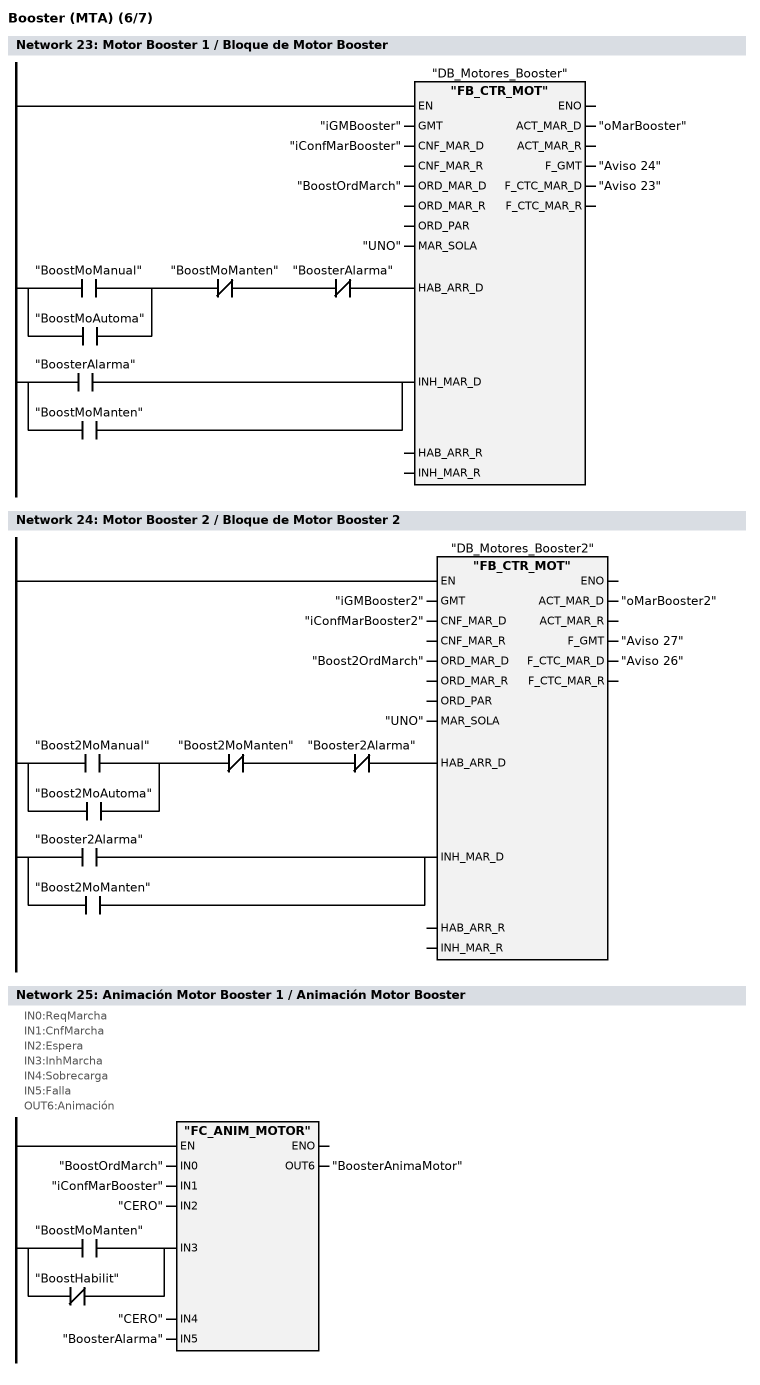
   RUNG wire#powerrail
      "DB_Motores_Booster"(HAB_ARR_D := wire#w2, INH_MAR_D := wire#w3, GMT := "iGMBooster", CNF_MAR_D := "iConfMarBooster", CNF_MAR_R :=, ORD_MAR_D := "BoostOrdMarch", ORD_MAR_R :=, ORD_PAR :=, MAR_SOLA := "UNO", HAB_ARR_R :=, INH_MAR_R :=, ACT_MAR_D => "oMarBooster", ACT_MAR_R =>, F_GMT => "Aviso 24", F_CTC_MAR_D => "Aviso 23", F_CTC_MAR_R =>)
   END_RUNG
   RUNG wire#powerrail
      Contact( "BoostMoManual" )
      wire#w1
      I_Contact( "BoostMoManten" )
      I_Contact( "BoosterAlarma" )
   END_RUNG wire#w2
   RUNG wire#powerrail
      Contact( "BoostMoAutoma" )
   END_RUNG wire#w1
   RUNG wire#powerrail
      Contact( "BoosterAlarma" )
   END_RUNG wire#w3
   RUNG wire#powerrail
      Contact( "BoostMoManten" )
   END_RUNG wire#w3
   // the same network as SCL:
   "DB_Motores_Booster"(GMT := "iGMBooster",   // "FB_CTR_MOT"
                        CNF_MAR_D := "iConfMarBooster",
                        ORD_MAR_D := "BoostOrdMarch",
                        MAR_SOLA := "UNO",
                        HAB_ARR_D := ("BoostMoManual" OR "BoostMoAutoma") AND NOT "BoostMoManten" AND NOT "BoosterAlarma",
                        INH_MAR_D := "BoosterAlarma" OR "BoostMoManten",
                        ACT_MAR_D => "oMarBooster",
                        F_GMT => "Aviso 24",
                        F_CTC_MAR_D => "Aviso 23");
END_REGION

REGION Network 24: Motor Booster 2 / Bloque de Motor Booster 2
   RUNG wire#powerrail
      "DB_Motores_Booster2"(HAB_ARR_D := wire#w2, INH_MAR_D := wire#w3, GMT := "iGMBooster2", CNF_MAR_D := "iConfMarBooster2", CNF_MAR_R :=, ORD_MAR_D := "Boost2OrdMarch", ORD_MAR_R :=, ORD_PAR :=, MAR_SOLA := "UNO", HAB_ARR_R :=, INH_MAR_R :=, ACT_MAR_D => "oMarBooster2", ACT_MAR_R =>, F_GMT => "Aviso 27", F_CTC_MAR_D => "Aviso 26", F_CTC_MAR_R =>)
   END_RUNG
   RUNG wire#powerrail
      Contact( "Boost2MoManual" )
      wire#w1
      I_Contact( "Boost2MoManten" )
      I_Contact( "Booster2Alarma" )
   END_RUNG wire#w2
   RUNG wire#powerrail
      Contact( "Boost2MoAutoma" )
   END_RUNG wire#w1
   RUNG wire#powerrail
      Contact( "Booster2Alarma" )
   END_RUNG wire#w3
   RUNG wire#powerrail
      Contact( "Boost2MoManten" )
   END_RUNG wire#w3
   // the same network as SCL:
   "DB_Motores_Booster2"(GMT := "iGMBooster2",   // "FB_CTR_MOT"
                         CNF_MAR_D := "iConfMarBooster2",
                         ORD_MAR_D := "Boost2OrdMarch",
                         MAR_SOLA := "UNO",
                         HAB_ARR_D := ("Boost2MoManual" OR "Boost2MoAutoma") AND NOT "Boost2MoManten" AND NOT "Booster2Alarma",
                         INH_MAR_D := "Booster2Alarma" OR "Boost2MoManten",
                         ACT_MAR_D => "oMarBooster2",
                         F_GMT => "Aviso 27",
                         F_CTC_MAR_D => "Aviso 26");
END_REGION

REGION Network 25: Animación Motor Booster 1 / Animación Motor Booster
   // IN0:ReqMarcha
   // IN1:CnfMarcha
   // IN2:Espera
   // IN3:InhMarcha
   // IN4:Sobrecarga
   // IN5:Falla
   // OUT6:Animación
   RUNG wire#powerrail
      "FC_ANIM_MOTOR"(IN0 := "BoostOrdMarch", IN1 := "iConfMarBooster", IN2 := "CERO", IN3 := wire#w1, IN4 := "CERO", IN5 := "BoosterAlarma", OUT6 => "BoosterAnimaMotor")
   END_RUNG
   RUNG wire#powerrail
      Contact( "BoostMoManten" )
   END_RUNG wire#w1
   RUNG wire#powerrail
      I_Contact( "BoostHabilit" )
   END_RUNG wire#w1
   // the same network as SCL:
   "FC_ANIM_MOTOR"(IN0 := "BoostOrdMarch",
                   IN1 := "iConfMarBooster",
                   IN2 := "CERO",
                   IN3 := "BoostMoManten" OR NOT "BoostHabilit",
                   IN4 := "CERO",
                   IN5 := "BoosterAlarma",
                   OUT6 => "BoosterAnimaMotor");
END_REGION

REGION Network 26: Animación Motor Booster 2
   // IN0:ReqMarcha
   // IN1:CnfMarcha
   // IN2:Espera
   // IN3:InhMarcha
   // IN4:Sobrecarga
   // IN5:Falla
   // OUT6:Animación
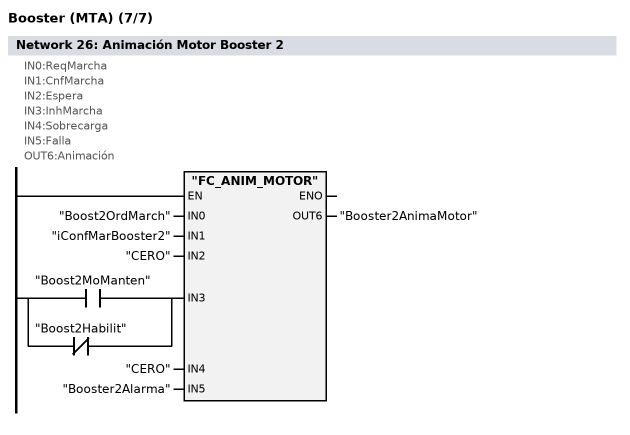
   RUNG wire#powerrail
      "FC_ANIM_MOTOR"(IN0 := "Boost2OrdMarch", IN1 := "iConfMarBooster2", IN2 := "CERO", IN3 := wire#w1, IN4 := "CERO", IN5 := "Booster2Alarma", OUT6 => "Booster2AnimaMotor")
   END_RUNG
   RUNG wire#powerrail
      Contact( "Boost2MoManten" )
   END_RUNG wire#w1
   RUNG wire#powerrail
      I_Contact( "Boost2Habilit" )
   END_RUNG wire#w1
   // the same network as SCL:
   "FC_ANIM_MOTOR"(IN0 := "Boost2OrdMarch",
                   IN1 := "iConfMarBooster2",
                   IN2 := "CERO",
                   IN3 := "Boost2MoManten" OR NOT "Boost2Habilit",
                   IN4 := "CERO",
                   IN5 := "Booster2Alarma",
                   OUT6 => "Booster2AnimaMotor");
END_REGION
END_FUNCTION

// folder: Compresores/Alta

FUNCTION "CompresoresAltaMTA" : Void   // FC13, LAD
{ S7_Optimized_Access := 'FALSE' }
VERSION : 0.1
BEGIN

REGION Network 1
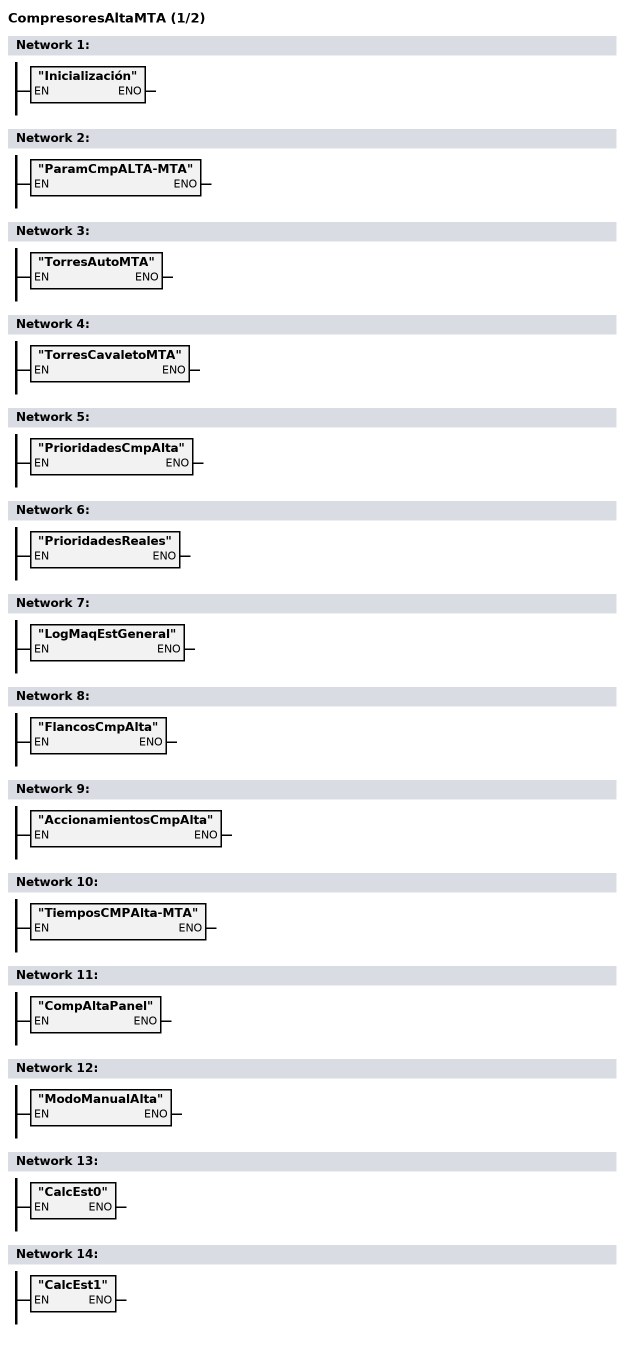
   RUNG wire#powerrail
      "Inicialización"()
   END_RUNG
   // the same network as SCL:
   "Inicialización"();
END_REGION

REGION Network 2
   RUNG wire#powerrail
      "ParamCmpALTA-MTA"()
   END_RUNG
   // the same network as SCL:
   "ParamCmpALTA-MTA"();
END_REGION

REGION Network 3
   RUNG wire#powerrail
      "TorresAutoMTA"()
   END_RUNG
   // the same network as SCL:
   "TorresAutoMTA"();
END_REGION

REGION Network 4
   RUNG wire#powerrail
      "TorresCavaletoMTA"()
   END_RUNG
   // the same network as SCL:
   "TorresCavaletoMTA"();
END_REGION

REGION Network 5
   RUNG wire#powerrail
      "PrioridadesCmpAlta"()
   END_RUNG
   // the same network as SCL:
   "PrioridadesCmpAlta"();
END_REGION

REGION Network 6
   RUNG wire#powerrail
      "PrioridadesReales"()
   END_RUNG
   // the same network as SCL:
   "PrioridadesReales"();
END_REGION

REGION Network 7
   RUNG wire#powerrail
      "LogMaqEstGeneral"()
   END_RUNG
   // the same network as SCL:
   "LogMaqEstGeneral"();
END_REGION

REGION Network 8
   RUNG wire#powerrail
      "FlancosCmpAlta"()
   END_RUNG
   // the same network as SCL:
   "FlancosCmpAlta"();
END_REGION

REGION Network 9
   RUNG wire#powerrail
      "AccionamientosCmpAlta"()
   END_RUNG
   // the same network as SCL:
   "AccionamientosCmpAlta"();
END_REGION

REGION Network 10
   RUNG wire#powerrail
      "TiemposCMPAlta-MTA"()
   END_RUNG
   // the same network as SCL:
   "TiemposCMPAlta-MTA"();
END_REGION

REGION Network 11
   RUNG wire#powerrail
      "CompAltaPanel"()
   END_RUNG
   // the same network as SCL:
   "CompAltaPanel"();
END_REGION

REGION Network 12
   RUNG wire#powerrail
      "ModoManualAlta"()
   END_RUNG
   // the same network as SCL:
   "ModoManualAlta"();
END_REGION

REGION Network 13
   RUNG wire#powerrail
      "CalcEst0"()
   END_RUNG
   // the same network as SCL:
   "CalcEst0"();
END_REGION

REGION Network 14
   RUNG wire#powerrail
      "CalcEst1"()
   END_RUNG
   // the same network as SCL:
   "CalcEst1"();
END_REGION

REGION Network 15
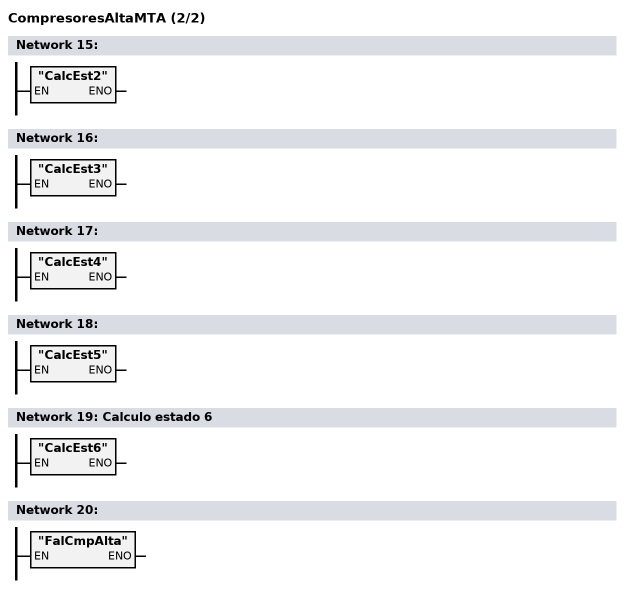
   RUNG wire#powerrail
      "CalcEst2"()
   END_RUNG
   // the same network as SCL:
   "CalcEst2"();
END_REGION

REGION Network 16
   RUNG wire#powerrail
      "CalcEst3"()
   END_RUNG
   // the same network as SCL:
   "CalcEst3"();
END_REGION

REGION Network 17
   RUNG wire#powerrail
      "CalcEst4"()
   END_RUNG
   // the same network as SCL:
   "CalcEst4"();
END_REGION

REGION Network 18
   RUNG wire#powerrail
      "CalcEst5"()
   END_RUNG
   // the same network as SCL:
   "CalcEst5"();
END_REGION

REGION Network 19: Calculo estado 6
   RUNG wire#powerrail
      "CalcEst6"()
   END_RUNG
   // the same network as SCL:
   "CalcEst6"();
END_REGION

REGION Network 20
   RUNG wire#powerrail
      "FalCmpAlta"()
   END_RUNG
   // the same network as SCL:
   "FalCmpAlta"();
END_REGION
END_FUNCTION

FUNCTION "ParamCmpALTA-MTA" : Void   // FC30, LAD
{ S7_Optimized_Access := 'FALSE' }
VERSION : 0.1
BEGIN

REGION Network 1
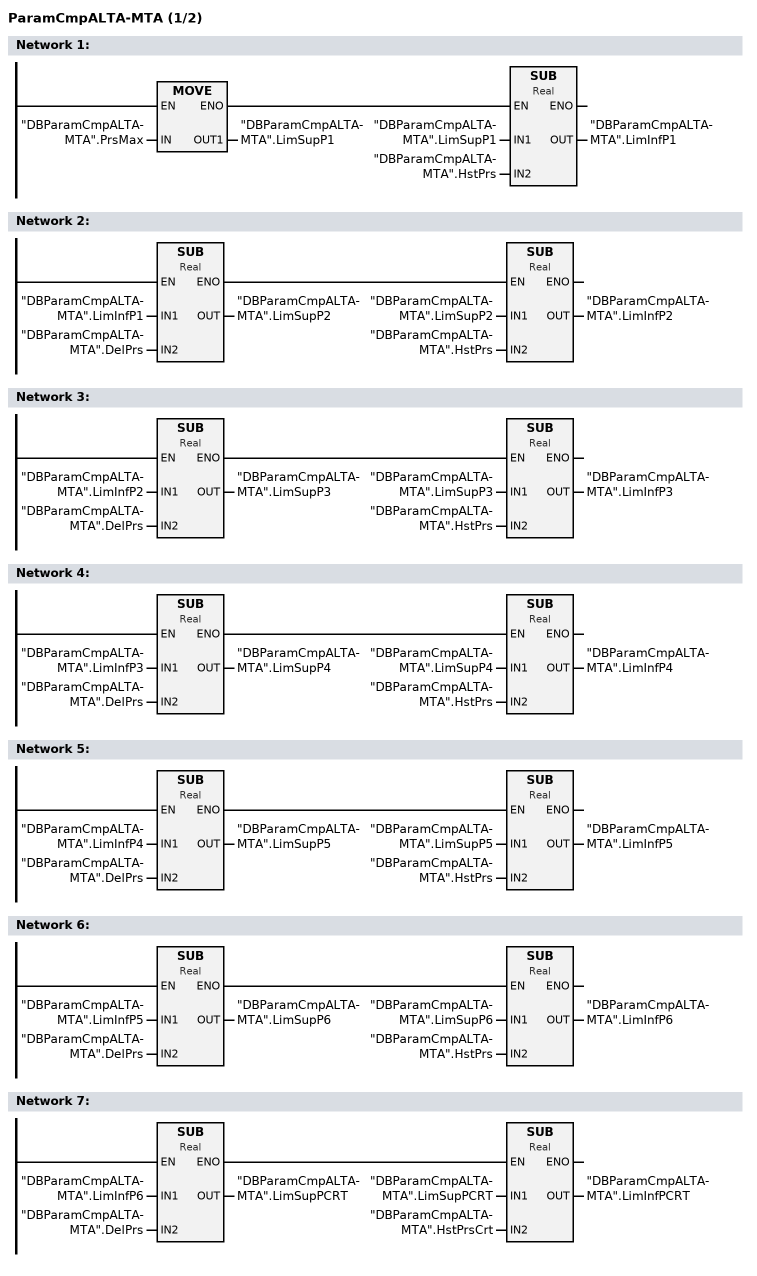
   RUNG wire#powerrail
      { S7_GenerateENO := "TRUE" } Move(in := "DBParamCmpALTA-MTA".PrsMax, out1 => "DBParamCmpALTA-MTA".LimSupP1)
      { S7_Templates := "SrcType := Real"; S7_GenerateENO := "TRUE" } Sub(in1 := "DBParamCmpALTA-MTA".LimSupP1, in2 := "DBParamCmpALTA-MTA".HstPrs, out => "DBParamCmpALTA-MTA".LimInfP1)
   END_RUNG
   // the same network as SCL:
   // ENO of a box is taken as its EN; it also drops when the box reports an error
   "DBParamCmpALTA-MTA".LimSupP1 := "DBParamCmpALTA-MTA".PrsMax;
   "DBParamCmpALTA-MTA".LimInfP1 := "DBParamCmpALTA-MTA".LimSupP1 - "DBParamCmpALTA-MTA".HstPrs;
END_REGION

REGION Network 2
   RUNG wire#powerrail
      { S7_Templates := "SrcType := Real"; S7_GenerateENO := "TRUE" } Sub(in1 := "DBParamCmpALTA-MTA".LimInfP1, in2 := "DBParamCmpALTA-MTA".DelPrs, out => "DBParamCmpALTA-MTA".LimSupP2)
      { S7_Templates := "SrcType := Real"; S7_GenerateENO := "TRUE" } Sub(in1 := "DBParamCmpALTA-MTA".LimSupP2, in2 := "DBParamCmpALTA-MTA".HstPrs, out => "DBParamCmpALTA-MTA".LimInfP2)
   END_RUNG
   // the same network as SCL:
   // ENO of a box is taken as its EN; it also drops when the box reports an error
   "DBParamCmpALTA-MTA".LimSupP2 := "DBParamCmpALTA-MTA".LimInfP1 - "DBParamCmpALTA-MTA".DelPrs;
   "DBParamCmpALTA-MTA".LimInfP2 := "DBParamCmpALTA-MTA".LimSupP2 - "DBParamCmpALTA-MTA".HstPrs;
END_REGION

REGION Network 3
   RUNG wire#powerrail
      { S7_Templates := "SrcType := Real"; S7_GenerateENO := "TRUE" } Sub(in1 := "DBParamCmpALTA-MTA".LimInfP2, in2 := "DBParamCmpALTA-MTA".DelPrs, out => "DBParamCmpALTA-MTA".LimSupP3)
      { S7_Templates := "SrcType := Real"; S7_GenerateENO := "TRUE" } Sub(in1 := "DBParamCmpALTA-MTA".LimSupP3, in2 := "DBParamCmpALTA-MTA".HstPrs, out => "DBParamCmpALTA-MTA".LimInfP3)
   END_RUNG
   // the same network as SCL:
   // ENO of a box is taken as its EN; it also drops when the box reports an error
   "DBParamCmpALTA-MTA".LimSupP3 := "DBParamCmpALTA-MTA".LimInfP2 - "DBParamCmpALTA-MTA".DelPrs;
   "DBParamCmpALTA-MTA".LimInfP3 := "DBParamCmpALTA-MTA".LimSupP3 - "DBParamCmpALTA-MTA".HstPrs;
END_REGION

REGION Network 4
   RUNG wire#powerrail
      { S7_Templates := "SrcType := Real"; S7_GenerateENO := "TRUE" } Sub(in1 := "DBParamCmpALTA-MTA".LimInfP3, in2 := "DBParamCmpALTA-MTA".DelPrs, out => "DBParamCmpALTA-MTA".LimSupP4)
      { S7_Templates := "SrcType := Real"; S7_GenerateENO := "TRUE" } Sub(in1 := "DBParamCmpALTA-MTA".LimSupP4, in2 := "DBParamCmpALTA-MTA".HstPrs, out => "DBParamCmpALTA-MTA".LimInfP4)
   END_RUNG
   // the same network as SCL:
   // ENO of a box is taken as its EN; it also drops when the box reports an error
   "DBParamCmpALTA-MTA".LimSupP4 := "DBParamCmpALTA-MTA".LimInfP3 - "DBParamCmpALTA-MTA".DelPrs;
   "DBParamCmpALTA-MTA".LimInfP4 := "DBParamCmpALTA-MTA".LimSupP4 - "DBParamCmpALTA-MTA".HstPrs;
END_REGION

REGION Network 5
   RUNG wire#powerrail
      { S7_Templates := "SrcType := Real"; S7_GenerateENO := "TRUE" } Sub(in1 := "DBParamCmpALTA-MTA".LimInfP4, in2 := "DBParamCmpALTA-MTA".DelPrs, out => "DBParamCmpALTA-MTA".LimSupP5)
      { S7_Templates := "SrcType := Real"; S7_GenerateENO := "TRUE" } Sub(in1 := "DBParamCmpALTA-MTA".LimSupP5, in2 := "DBParamCmpALTA-MTA".HstPrs, out => "DBParamCmpALTA-MTA".LimInfP5)
   END_RUNG
   // the same network as SCL:
   // ENO of a box is taken as its EN; it also drops when the box reports an error
   "DBParamCmpALTA-MTA".LimSupP5 := "DBParamCmpALTA-MTA".LimInfP4 - "DBParamCmpALTA-MTA".DelPrs;
   "DBParamCmpALTA-MTA".LimInfP5 := "DBParamCmpALTA-MTA".LimSupP5 - "DBParamCmpALTA-MTA".HstPrs;
END_REGION

REGION Network 6
   RUNG wire#powerrail
      { S7_Templates := "SrcType := Real"; S7_GenerateENO := "TRUE" } Sub(in1 := "DBParamCmpALTA-MTA".LimInfP5, in2 := "DBParamCmpALTA-MTA".DelPrs, out => "DBParamCmpALTA-MTA".LimSupP6)
      { S7_Templates := "SrcType := Real"; S7_GenerateENO := "TRUE" } Sub(in1 := "DBParamCmpALTA-MTA".LimSupP6, in2 := "DBParamCmpALTA-MTA".HstPrs, out => "DBParamCmpALTA-MTA".LimInfP6)
   END_RUNG
   // the same network as SCL:
   // ENO of a box is taken as its EN; it also drops when the box reports an error
   "DBParamCmpALTA-MTA".LimSupP6 := "DBParamCmpALTA-MTA".LimInfP5 - "DBParamCmpALTA-MTA".DelPrs;
   "DBParamCmpALTA-MTA".LimInfP6 := "DBParamCmpALTA-MTA".LimSupP6 - "DBParamCmpALTA-MTA".HstPrs;
END_REGION

REGION Network 7
   RUNG wire#powerrail
      { S7_Templates := "SrcType := Real"; S7_GenerateENO := "TRUE" } Sub(in1 := "DBParamCmpALTA-MTA".LimInfP6, in2 := "DBParamCmpALTA-MTA".DelPrs, out => "DBParamCmpALTA-MTA".LimSupPCRT)
      { S7_Templates := "SrcType := Real"; S7_GenerateENO := "TRUE" } Sub(in1 := "DBParamCmpALTA-MTA".LimSupPCRT, in2 := "DBParamCmpALTA-MTA".HstPrsCrt, out => "DBParamCmpALTA-MTA".LimInfPCRT)
   END_RUNG
   // the same network as SCL:
   // ENO of a box is taken as its EN; it also drops when the box reports an error
   "DBParamCmpALTA-MTA".LimSupPCRT := "DBParamCmpALTA-MTA".LimInfP6 - "DBParamCmpALTA-MTA".DelPrs;
   "DBParamCmpALTA-MTA".LimInfPCRT := "DBParamCmpALTA-MTA".LimSupPCRT - "DBParamCmpALTA-MTA".HstPrsCrt;
END_REGION

REGION Network 8: Falla General Flujostato Cavaleto
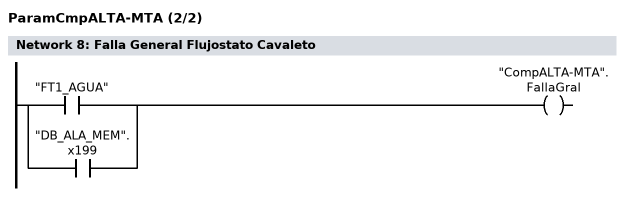
   RUNG wire#powerrail
      Contact( "FT1_AGUA" )
      wire#w1
      Coil( "CompALTA-MTA".FallaGral )
   END_RUNG
   RUNG wire#powerrail
      Contact( "DB_ALA_MEM".x199 )
   END_RUNG wire#w1
   // the same network as SCL:
   "CompALTA-MTA".FallaGral := "FT1_AGUA" OR "DB_ALA_MEM".x199;
END_REGION
END_FUNCTION

FUNCTION "TiemposCMPAlta-MTA" : Void   // FC31, LAD
{ S7_Optimized_Access := 'FALSE' }
VERSION : 0.1
   VAR_TEMP   // added for the SCL form of the ladder/FBD networks
      _s5time1 : S5Time;
   END_VAR
BEGIN

REGION Network 1
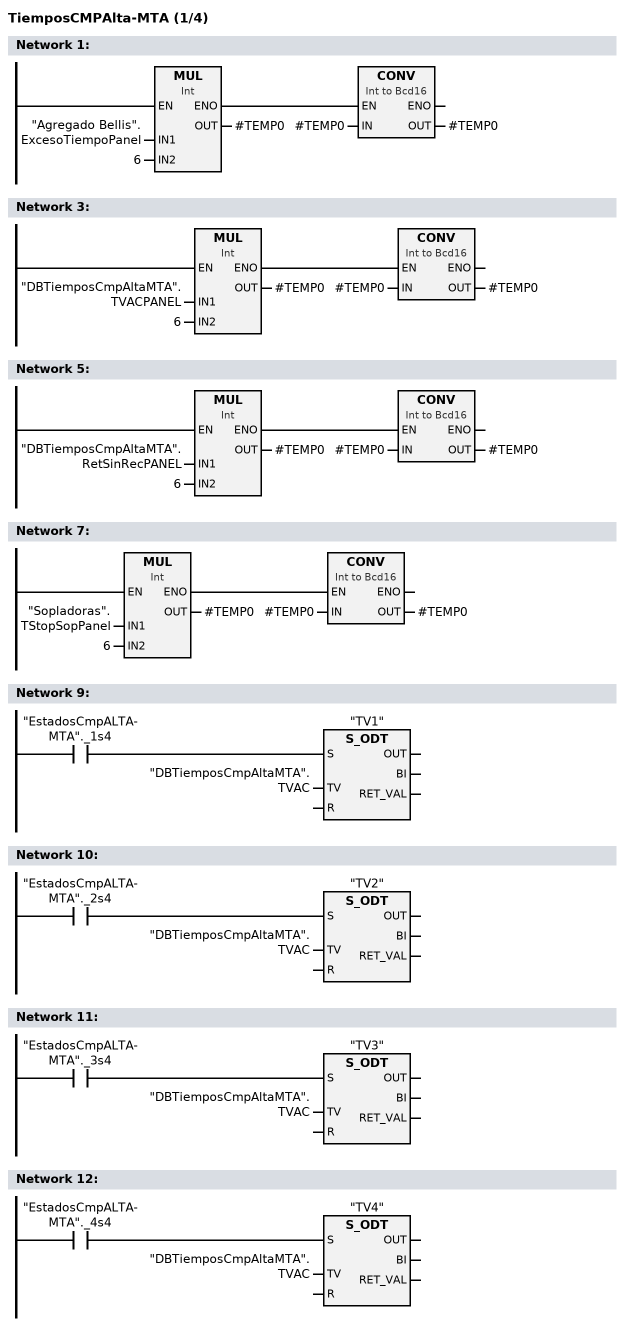
   RUNG wire#powerrail
      { S7_Templates := "SrcType := Int"; S7_GenerateENO := "TRUE" } Mul(in1 := "Agregado Bellis".ExcesoTiempoPanel, in2 := 6, out => #TEMP0)
      { S7_Templates := "[SrcType := Int, DestType := Bcd16]"; S7_GenerateENO := "TRUE" } Convert(in := #TEMP0, out => #TEMP0)
   END_RUNG
   // the same network as SCL:
   // ENO of a box is taken as its EN; it also drops when the box reports an error
   #TEMP0 := "Agregado Bellis".ExcesoTiempoPanel * 6;
   #TEMP0 := INT_TO_BCD16(#TEMP0);
END_REGION

REGION Network 2 (STL)
         L     12288;
         L     #TEMP0;
         OW;
         T     "Agregado Bellis".ExcesoTiempo;
         NOP   0;
END_REGION

REGION Network 3
   RUNG wire#powerrail
      { S7_Templates := "SrcType := Int"; S7_GenerateENO := "TRUE" } Mul(in1 := "DBTiemposCmpAltaMTA".TVACPANEL, in2 := 6, out => #TEMP0)
      { S7_Templates := "[SrcType := Int, DestType := Bcd16]"; S7_GenerateENO := "TRUE" } Convert(in := #TEMP0, out => #TEMP0)
   END_RUNG
   // the same network as SCL:
   // ENO of a box is taken as its EN; it also drops when the box reports an error
   #TEMP0 := "DBTiemposCmpAltaMTA".TVACPANEL * 6;
   #TEMP0 := INT_TO_BCD16(#TEMP0);
END_REGION

REGION Network 4 (STL)
         L     12288;
         L     #TEMP0;
         OW;
         T     "DBTiemposCmpAltaMTA".TVAC;
         NOP   0;
END_REGION

REGION Network 5
   RUNG wire#powerrail
      { S7_Templates := "SrcType := Int"; S7_GenerateENO := "TRUE" } Mul(in1 := "DBTiemposCmpAltaMTA".RetSinRecPANEL, in2 := 6, out => #TEMP0)
      { S7_Templates := "[SrcType := Int, DestType := Bcd16]"; S7_GenerateENO := "TRUE" } Convert(in := #TEMP0, out => #TEMP0)
   END_RUNG
   // the same network as SCL:
   // ENO of a box is taken as its EN; it also drops when the box reports an error
   #TEMP0 := "DBTiemposCmpAltaMTA".RetSinRecPANEL * 6;
   #TEMP0 := INT_TO_BCD16(#TEMP0);
END_REGION

REGION Network 6 (STL)
         L     12288;
         L     #TEMP0;
         OW;
         T     "DBTiemposCmpAltaMTA".RetSinRec;
         NOP   0;
END_REGION

REGION Network 7
   RUNG wire#powerrail
      { S7_Templates := "SrcType := Int"; S7_GenerateENO := "TRUE" } Mul(in1 := "Sopladoras".TStopSopPanel, in2 := 6, out => #TEMP0)
      { S7_Templates := "[SrcType := Int, DestType := Bcd16]"; S7_GenerateENO := "TRUE" } Convert(in := #TEMP0, out => #TEMP0)
   END_RUNG
   // the same network as SCL:
   // ENO of a box is taken as its EN; it also drops when the box reports an error
   #TEMP0 := "Sopladoras".TStopSopPanel * 6;
   #TEMP0 := INT_TO_BCD16(#TEMP0);
END_REGION

REGION Network 8 (STL)
         L     12288;
         L     #TEMP0;
         OW;
         T     "Sopladoras".TStopSop;
         NOP   0;
END_REGION

REGION Network 9
   RUNG wire#powerrail
      Contact( "EstadosCmpALTA-MTA"._1s4 )
      S_ODT(T_NO := "TV1", TV := "DBTiemposCmpAltaMTA".TVAC, R :=, BI =>, RET_VAL =>)
   END_RUNG
   // the same network as SCL:
   #_s5time1 := S_ODT(T_NO := "TV1", S := "EstadosCmpALTA-MTA"._1s4, TV := "DBTiemposCmpAltaMTA".TVAC);
END_REGION

REGION Network 10
   RUNG wire#powerrail
      Contact( "EstadosCmpALTA-MTA"._2s4 )
      S_ODT(T_NO := "TV2", TV := "DBTiemposCmpAltaMTA".TVAC, R :=, BI =>, RET_VAL =>)
   END_RUNG
   // the same network as SCL:
   #_s5time1 := S_ODT(T_NO := "TV2", S := "EstadosCmpALTA-MTA"._2s4, TV := "DBTiemposCmpAltaMTA".TVAC);
END_REGION

REGION Network 11
   RUNG wire#powerrail
      Contact( "EstadosCmpALTA-MTA"._3s4 )
      S_ODT(T_NO := "TV3", TV := "DBTiemposCmpAltaMTA".TVAC, R :=, BI =>, RET_VAL =>)
   END_RUNG
   // the same network as SCL:
   #_s5time1 := S_ODT(T_NO := "TV3", S := "EstadosCmpALTA-MTA"._3s4, TV := "DBTiemposCmpAltaMTA".TVAC);
END_REGION

REGION Network 12
   RUNG wire#powerrail
      Contact( "EstadosCmpALTA-MTA"._4s4 )
      S_ODT(T_NO := "TV4", TV := "DBTiemposCmpAltaMTA".TVAC, R :=, BI =>, RET_VAL =>)
   END_RUNG
   // the same network as SCL:
   #_s5time1 := S_ODT(T_NO := "TV4", S := "EstadosCmpALTA-MTA"._4s4, TV := "DBTiemposCmpAltaMTA".TVAC);
END_REGION

REGION Network 13
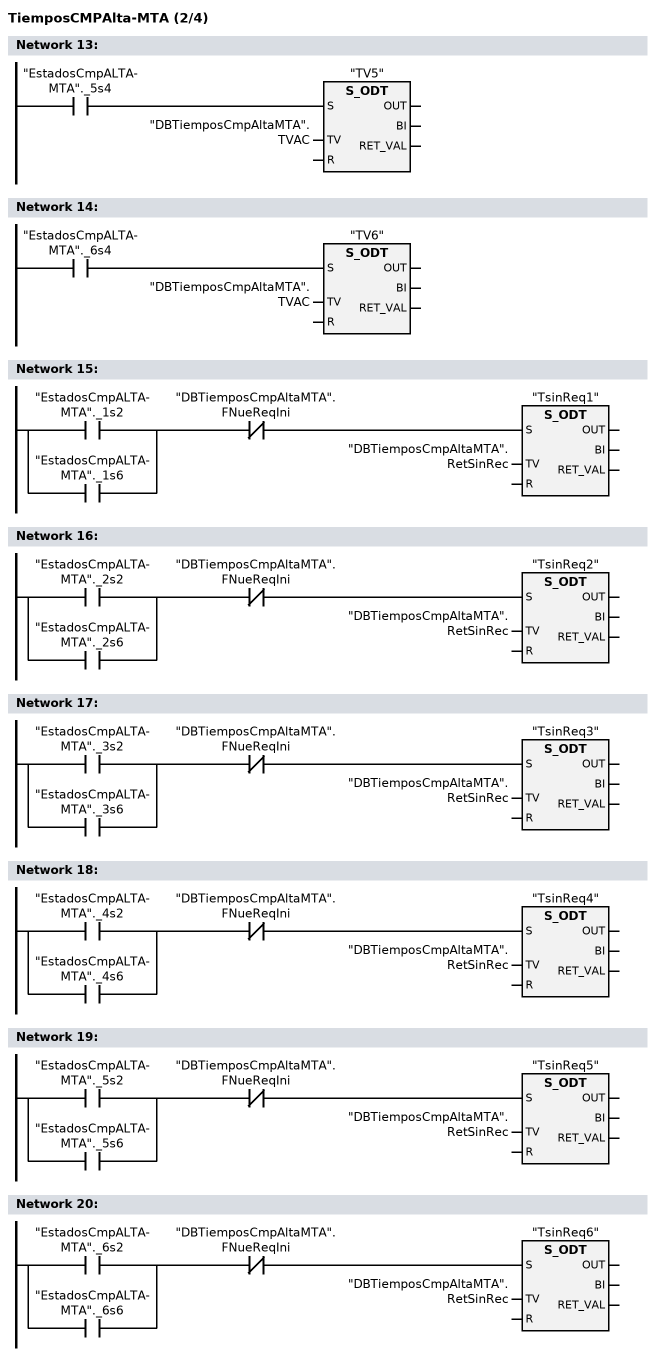
   RUNG wire#powerrail
      Contact( "EstadosCmpALTA-MTA"._5s4 )
      S_ODT(T_NO := "TV5", TV := "DBTiemposCmpAltaMTA".TVAC, R :=, BI =>, RET_VAL =>)
   END_RUNG
   // the same network as SCL:
   #_s5time1 := S_ODT(T_NO := "TV5", S := "EstadosCmpALTA-MTA"._5s4, TV := "DBTiemposCmpAltaMTA".TVAC);
END_REGION

REGION Network 14
   RUNG wire#powerrail
      Contact( "EstadosCmpALTA-MTA"._6s4 )
      S_ODT(T_NO := "TV6", TV := "DBTiemposCmpAltaMTA".TVAC, R :=, BI =>, RET_VAL =>)
   END_RUNG
   // the same network as SCL:
   #_s5time1 := S_ODT(T_NO := "TV6", S := "EstadosCmpALTA-MTA"._6s4, TV := "DBTiemposCmpAltaMTA".TVAC);
END_REGION

REGION Network 15
   RUNG wire#powerrail
      Contact( "EstadosCmpALTA-MTA"._1s2 )
      wire#w1
      I_Contact( "DBTiemposCmpAltaMTA".FNueReqIni )
      S_ODT(T_NO := "TsinReq1", TV := "DBTiemposCmpAltaMTA".RetSinRec, R :=, BI =>, RET_VAL =>)
   END_RUNG
   RUNG wire#powerrail
      Contact( "EstadosCmpALTA-MTA"._1s6 )
   END_RUNG wire#w1
   // the same network as SCL:
   #_s5time1 := S_ODT(T_NO := "TsinReq1",
                      S := ("EstadosCmpALTA-MTA"._1s2 OR "EstadosCmpALTA-MTA"._1s6) AND NOT "DBTiemposCmpAltaMTA".FNueReqIni,
                      TV := "DBTiemposCmpAltaMTA".RetSinRec);
END_REGION

REGION Network 16
   RUNG wire#powerrail
      Contact( "EstadosCmpALTA-MTA"._2s2 )
      wire#w1
      I_Contact( "DBTiemposCmpAltaMTA".FNueReqIni )
      S_ODT(T_NO := "TsinReq2", TV := "DBTiemposCmpAltaMTA".RetSinRec, R :=, BI =>, RET_VAL =>)
   END_RUNG
   RUNG wire#powerrail
      Contact( "EstadosCmpALTA-MTA"._2s6 )
   END_RUNG wire#w1
   // the same network as SCL:
   #_s5time1 := S_ODT(T_NO := "TsinReq2",
                      S := ("EstadosCmpALTA-MTA"._2s2 OR "EstadosCmpALTA-MTA"._2s6) AND NOT "DBTiemposCmpAltaMTA".FNueReqIni,
                      TV := "DBTiemposCmpAltaMTA".RetSinRec);
END_REGION

REGION Network 17
   RUNG wire#powerrail
      Contact( "EstadosCmpALTA-MTA"._3s2 )
      wire#w1
      I_Contact( "DBTiemposCmpAltaMTA".FNueReqIni )
      S_ODT(T_NO := "TsinReq3", TV := "DBTiemposCmpAltaMTA".RetSinRec, R :=, BI =>, RET_VAL =>)
   END_RUNG
   RUNG wire#powerrail
      Contact( "EstadosCmpALTA-MTA"._3s6 )
   END_RUNG wire#w1
   // the same network as SCL:
   #_s5time1 := S_ODT(T_NO := "TsinReq3",
                      S := ("EstadosCmpALTA-MTA"._3s2 OR "EstadosCmpALTA-MTA"._3s6) AND NOT "DBTiemposCmpAltaMTA".FNueReqIni,
                      TV := "DBTiemposCmpAltaMTA".RetSinRec);
END_REGION

REGION Network 18
   RUNG wire#powerrail
      Contact( "EstadosCmpALTA-MTA"._4s2 )
      wire#w1
      I_Contact( "DBTiemposCmpAltaMTA".FNueReqIni )
      S_ODT(T_NO := "TsinReq4", TV := "DBTiemposCmpAltaMTA".RetSinRec, R :=, BI =>, RET_VAL =>)
   END_RUNG
   RUNG wire#powerrail
      Contact( "EstadosCmpALTA-MTA"._4s6 )
   END_RUNG wire#w1
   // the same network as SCL:
   #_s5time1 := S_ODT(T_NO := "TsinReq4",
                      S := ("EstadosCmpALTA-MTA"._4s2 OR "EstadosCmpALTA-MTA"._4s6) AND NOT "DBTiemposCmpAltaMTA".FNueReqIni,
                      TV := "DBTiemposCmpAltaMTA".RetSinRec);
END_REGION

REGION Network 19
   RUNG wire#powerrail
      Contact( "EstadosCmpALTA-MTA"._5s2 )
      wire#w1
      I_Contact( "DBTiemposCmpAltaMTA".FNueReqIni )
      S_ODT(T_NO := "TsinReq5", TV := "DBTiemposCmpAltaMTA".RetSinRec, R :=, BI =>, RET_VAL =>)
   END_RUNG
   RUNG wire#powerrail
      Contact( "EstadosCmpALTA-MTA"._5s6 )
   END_RUNG wire#w1
   // the same network as SCL:
   #_s5time1 := S_ODT(T_NO := "TsinReq5",
                      S := ("EstadosCmpALTA-MTA"._5s2 OR "EstadosCmpALTA-MTA"._5s6) AND NOT "DBTiemposCmpAltaMTA".FNueReqIni,
                      TV := "DBTiemposCmpAltaMTA".RetSinRec);
END_REGION

REGION Network 20
   RUNG wire#powerrail
      Contact( "EstadosCmpALTA-MTA"._6s2 )
      wire#w1
      I_Contact( "DBTiemposCmpAltaMTA".FNueReqIni )
      S_ODT(T_NO := "TsinReq6", TV := "DBTiemposCmpAltaMTA".RetSinRec, R :=, BI =>, RET_VAL =>)
   END_RUNG
   RUNG wire#powerrail
      Contact( "EstadosCmpALTA-MTA"._6s6 )
   END_RUNG wire#w1
   // the same network as SCL:
   #_s5time1 := S_ODT(T_NO := "TsinReq6",
                      S := ("EstadosCmpALTA-MTA"._6s2 OR "EstadosCmpALTA-MTA"._6s6) AND NOT "DBTiemposCmpAltaMTA".FNueReqIni,
                      TV := "DBTiemposCmpAltaMTA".RetSinRec);
END_REGION

REGION Network 21
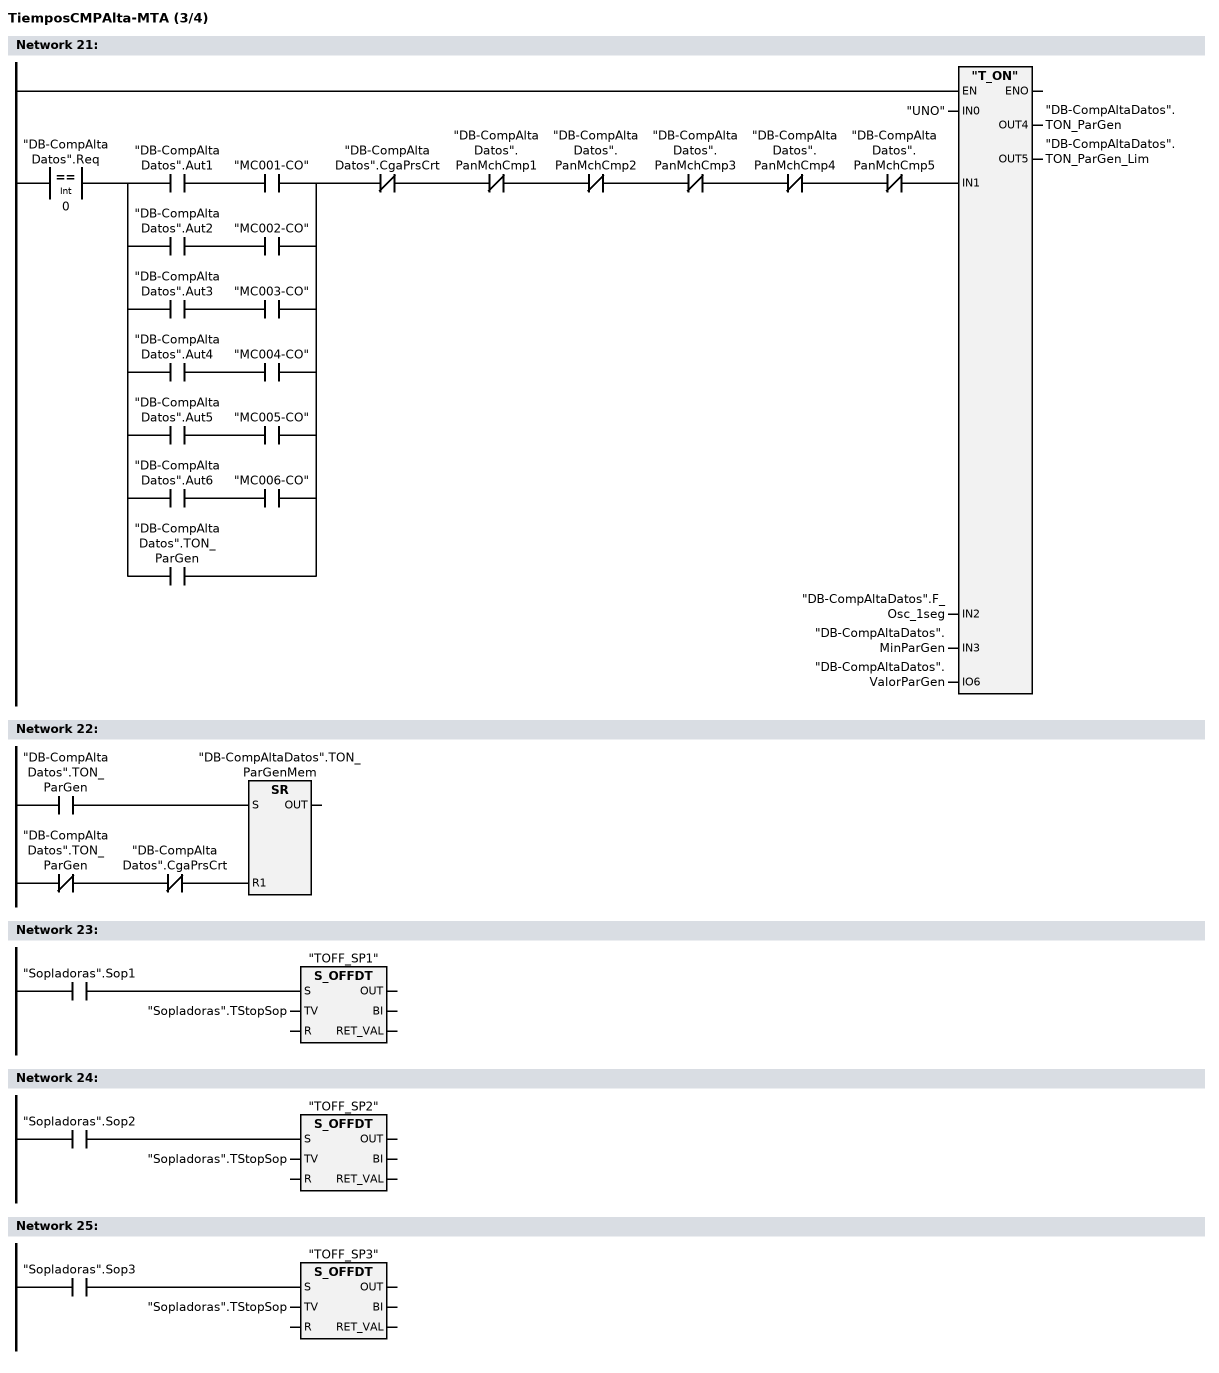
   RUNG wire#powerrail
      "T_ON"(IN1 := wire#w3, IN0 := "UNO", IN2 := "DB-CompAltaDatos".F_Osc_1seg, IN3 := "DB-CompAltaDatos".MinParGen, IO6 := "DB-CompAltaDatos".ValorParGen, OUT4 => "DB-CompAltaDatos".TON_ParGen, OUT5 => "DB-CompAltaDatos".TON_ParGen_Lim)
   END_RUNG
   RUNG wire#powerrail
      { S7_Templates := "SrcType := Int" } EQ_Contact(in1 := "DB-CompAltaDatos".Req, in2 := 0)
      wire#w1
      Contact( "DB-CompAltaDatos".Aut1 )
      Contact( "MC001-CO" )
      wire#w2
      I_Contact( "DB-CompAltaDatos".CgaPrsCrt )
      I_Contact( "DB-CompAltaDatos".PanMchCmp1 )
      I_Contact( "DB-CompAltaDatos".PanMchCmp2 )
      I_Contact( "DB-CompAltaDatos".PanMchCmp3 )
      I_Contact( "DB-CompAltaDatos".PanMchCmp4 )
      I_Contact( "DB-CompAltaDatos".PanMchCmp5 )
   END_RUNG wire#w3
   RUNG wire#w1
      Contact( "DB-CompAltaDatos".Aut2 )
      Contact( "MC002-CO" )
   END_RUNG wire#w2
   RUNG wire#w1
      Contact( "DB-CompAltaDatos".Aut3 )
      Contact( "MC003-CO" )
   END_RUNG wire#w2
   RUNG wire#w1
      Contact( "DB-CompAltaDatos".Aut4 )
      Contact( "MC004-CO" )